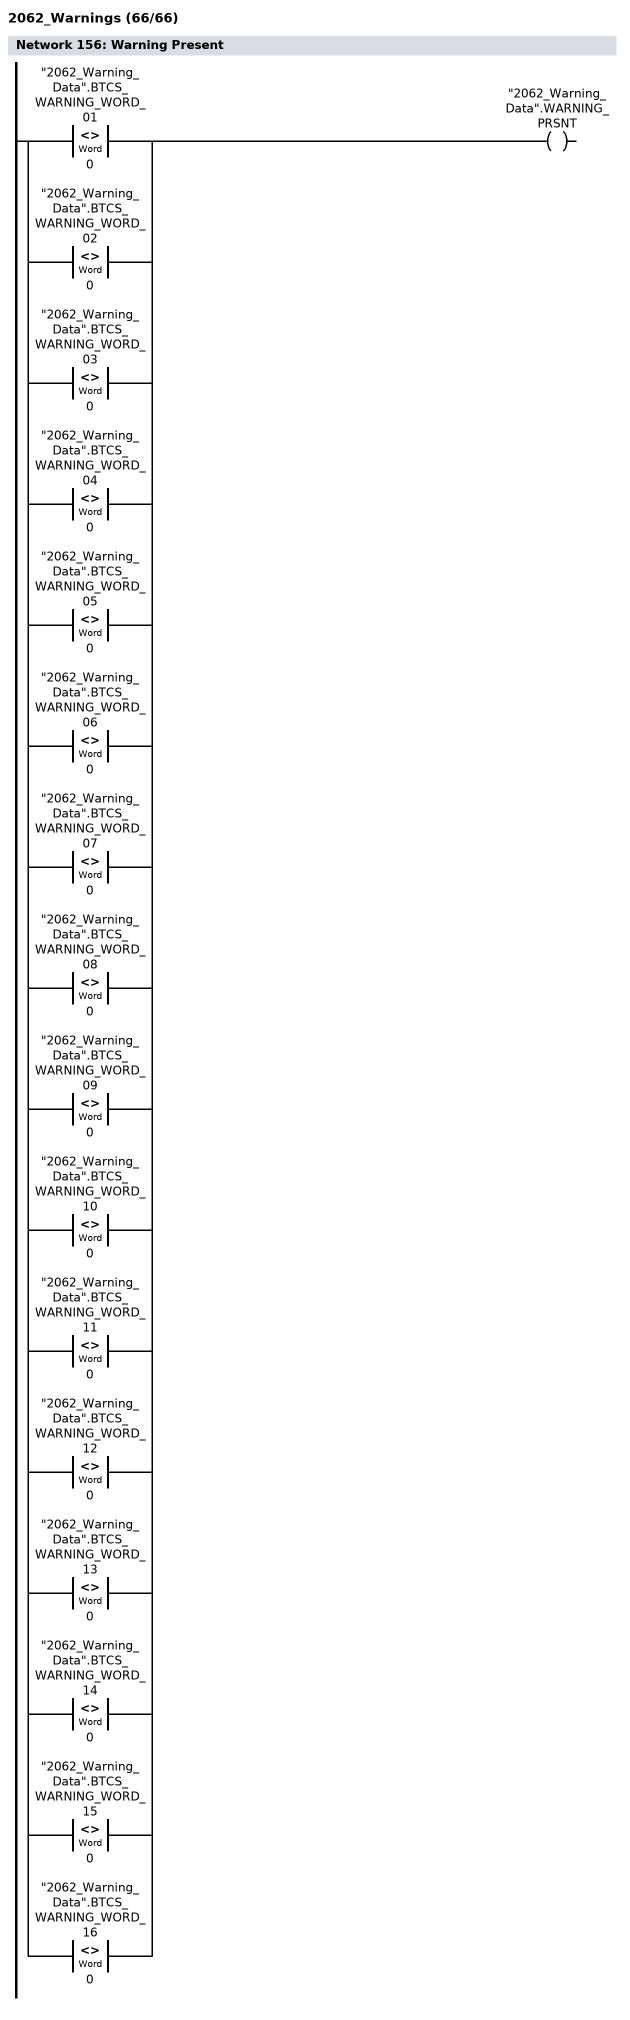
   RUNG wire#powerrail
      { S7_Templates := "SrcType := Word" } NE_Contact(in1 := "2062_Warning_Data".BTCS_WARNING_WORD_01, in2 := 0)
      wire#w1
      Coil( "2062_Warning_Data".WARNING_PRSNT )
   END_RUNG
   RUNG wire#powerrail
      { S7_Templates := "SrcType := Word" } NE_Contact(in1 := "2062_Warning_Data".BTCS_WARNING_WORD_02, in2 := 0)
   END_RUNG wire#w1
   RUNG wire#powerrail
      { S7_Templates := "SrcType := Word" } NE_Contact(in1 := "2062_Warning_Data".BTCS_WARNING_WORD_03, in2 := 0)
   END_RUNG wire#w1
   RUNG wire#powerrail
      { S7_Templates := "SrcType := Word" } NE_Contact(in1 := "2062_Warning_Data".BTCS_WARNING_WORD_04, in2 := 0)
   END_RUNG wire#w1
   RUNG wire#powerrail
      { S7_Templates := "SrcType := Word" } NE_Contact(in1 := "2062_Warning_Data".BTCS_WARNING_WORD_05, in2 := 0)
   END_RUNG wire#w1
   RUNG wire#powerrail
      { S7_Templates := "SrcType := Word" } NE_Contact(in1 := "2062_Warning_Data".BTCS_WARNING_WORD_06, in2 := 0)
   END_RUNG wire#w1
   RUNG wire#powerrail
      { S7_Templates := "SrcType := Word" } NE_Contact(in1 := "2062_Warning_Data".BTCS_WARNING_WORD_07, in2 := 0)
   END_RUNG wire#w1
   RUNG wire#powerrail
      { S7_Templates := "SrcType := Word" } NE_Contact(in1 := "2062_Warning_Data".BTCS_WARNING_WORD_08, in2 := 0)
   END_RUNG wire#w1
   RUNG wire#powerrail
      { S7_Templates := "SrcType := Word" } NE_Contact(in1 := "2062_Warning_Data".BTCS_WARNING_WORD_09, in2 := 0)
   END_RUNG wire#w1
   RUNG wire#powerrail
      { S7_Templates := "SrcType := Word" } NE_Contact(in1 := "2062_Warning_Data".BTCS_WARNING_WORD_10, in2 := 0)
   END_RUNG wire#w1
   RUNG wire#powerrail
      { S7_Templates := "SrcType := Word" } NE_Contact(in1 := "2062_Warning_Data".BTCS_WARNING_WORD_11, in2 := 0)
   END_RUNG wire#w1
   RUNG wire#powerrail
      { S7_Templates := "SrcType := Word" } NE_Contact(in1 := "2062_Warning_Data".BTCS_WARNING_WORD_12, in2 := 0)
   END_RUNG wire#w1
   RUNG wire#powerrail
      { S7_Templates := "SrcType := Word" } NE_Contact(in1 := "2062_Warning_Data".BTCS_WARNING_WORD_13, in2 := 0)
   END_RUNG wire#w1
   RUNG wire#powerrail
      { S7_Templates := "SrcType := Word" } NE_Contact(in1 := "2062_Warning_Data".BTCS_WARNING_WORD_14, in2 := 0)
   END_RUNG wire#w1
   RUNG wire#powerrail
      { S7_Templates := "SrcType := Word" } NE_Contact(in1 := "2062_Warning_Data".BTCS_WARNING_WORD_15, in2 := 0)
   END_RUNG wire#w1
   RUNG wire#powerrail
      { S7_Templates := "SrcType := Word" } NE_Contact(in1 := "2062_Warning_Data".BTCS_WARNING_WORD_16, in2 := 0)
   END_RUNG wire#w1
   // the same network as SCL:
   "2062_Warning_Data".WARNING_PRSNT := ("2062_Warning_Data".BTCS_WARNING_WORD_01 <> 0) OR ("2062_Warning_Data".BTCS_WARNING_WORD_02 <> 0) OR ("2062_Warning_Data".BTCS_WARNING_WORD_03 <> 0) OR ("2062_Warning_Data".BTCS_WARNING_WORD_04 <> 0) OR ("2062_Warning_Data".BTCS_WARNING_WORD_05 <> 0) OR ("2062_Warning_Data".BTCS_WARNING_WORD_06 <> 0) OR ("2062_Warning_Data".BTCS_WARNING_WORD_07 <> 0) OR ("2062_Warning_Data".BTCS_WARNING_WORD_08 <> 0) OR ("2062_Warning_Data".BTCS_WARNING_WORD_09 <> 0) OR ("2062_Warning_Data".BTCS_WARNING_WORD_10 <> 0) OR ("2062_Warning_Data".BTCS_WARNING_WORD_11 <> 0) OR ("2062_Warning_Data".BTCS_WARNING_WORD_12 <> 0) OR ("2062_Warning_Data".BTCS_WARNING_WORD_13 <> 0) OR ("2062_Warning_Data".BTCS_WARNING_WORD_14 <> 0) OR ("2062_Warning_Data".BTCS_WARNING_WORD_15 <> 0) OR ("2062_Warning_Data".BTCS_WARNING_WORD_16 <> 0);
END_REGION
END_FUNCTION

FUNCTION "2068_Sys_Status" : Void   // FC2068, LAD
TITLE = System Status
{ S7_Optimized_Access := 'TRUE' }
AUTHOR : JRS
VERSION : 0.1
// For the determination of specific system status information as required by the code
   VAR_TEMP
      RET_VAL_1 : Int;
      LOCAL_DATE_AND_TIME : DTL;
   END_VAR
   VAR_TEMP   // added for the SCL form of the ladder/FBD networks
      _w1 : Bool;
      _w2 : Bool;
      _w3 : Bool;
      _w4 : Bool;
   END_VAR
BEGIN

REGION Network 1: Port GTT Open Timer For Flow De-Bounce
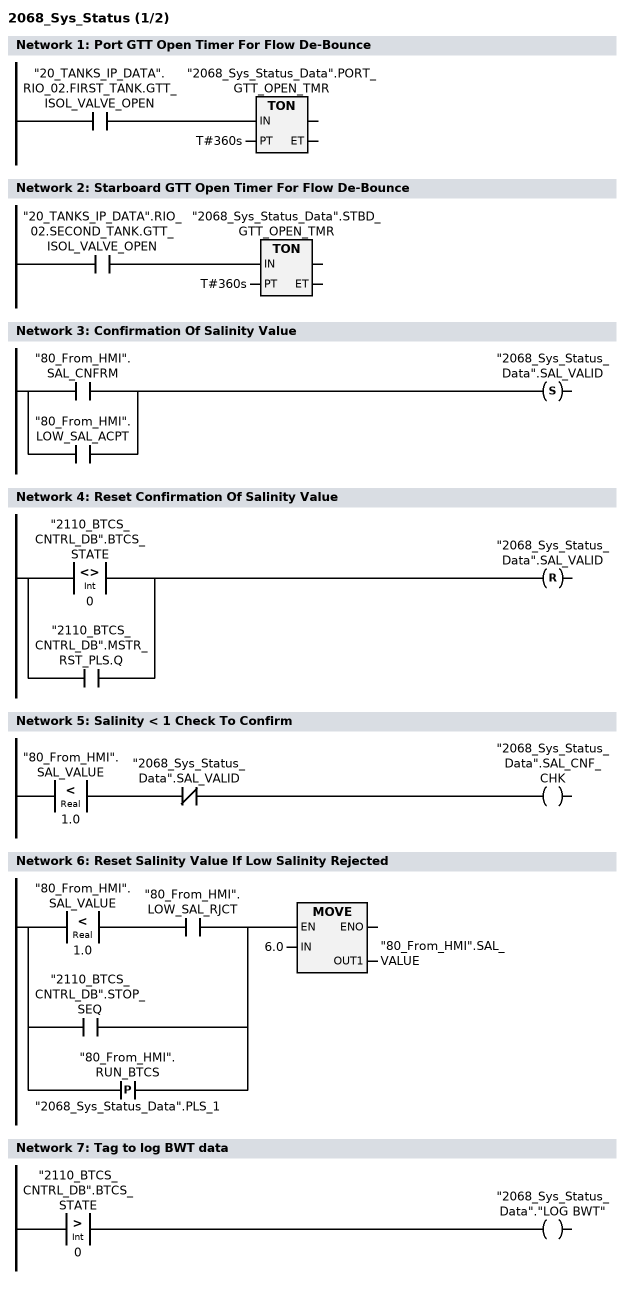
   "2068_Sys_Status_Data".PORT_GTT_OPEN_TMR.TON(IN := "20_TANKS_IP_DATA".RIO_02.FIRST_TANK.GTT_ISOL_VALVE_OPEN,
                           PT := T#360s);
END_REGION

REGION Network 2: Starboard GTT Open Timer For Flow De-Bounce
   "2068_Sys_Status_Data".STBD_GTT_OPEN_TMR.TON(IN := "20_TANKS_IP_DATA".RIO_02.SECOND_TANK.GTT_ISOL_VALVE_OPEN,
                           PT := T#360s);
END_REGION

REGION Network 3: Confirmation Of Salinity Value
   RUNG wire#powerrail
      Contact( "80_From_HMI".SAL_CNFRM )
      wire#w1
      S_Coil( "2068_Sys_Status_Data".SAL_VALID )
   END_RUNG
   RUNG wire#powerrail
      Contact( "80_From_HMI".LOW_SAL_ACPT )
   END_RUNG wire#w1
   // the same network as SCL:
   IF "80_From_HMI".SAL_CNFRM OR "80_From_HMI".LOW_SAL_ACPT THEN
       "2068_Sys_Status_Data".SAL_VALID := TRUE;
   END_IF;
END_REGION

REGION Network 4: Reset Confirmation Of Salinity Value
   RUNG wire#powerrail
      { S7_Templates := "SrcType := Int" } NE_Contact(in1 := "2110_BTCS_CNTRL_DB".BTCS_STATE, in2 := 0)
      wire#w1
      R_Coil( "2068_Sys_Status_Data".SAL_VALID )
   END_RUNG
   RUNG wire#powerrail
      Contact( "2110_BTCS_CNTRL_DB".MSTR_RST_PLS.Q )
   END_RUNG wire#w1
   // the same network as SCL:
   IF ("2110_BTCS_CNTRL_DB".BTCS_STATE <> 0) OR "2110_BTCS_CNTRL_DB".MSTR_RST_PLS.Q THEN
       "2068_Sys_Status_Data".SAL_VALID := FALSE;
   END_IF;
END_REGION

REGION Network 5: Salinity < 1 Check To Confirm
   RUNG wire#powerrail
      { S7_Templates := "SrcType := Real" } LT_Contact(in1 := "80_From_HMI".SAL_VALUE, in2 := 1.0)
      I_Contact( "2068_Sys_Status_Data".SAL_VALID )
      Coil( "2068_Sys_Status_Data".SAL_CNF_CHK )
   END_RUNG
   // the same network as SCL:
   "2068_Sys_Status_Data".SAL_CNF_CHK := ("80_From_HMI".SAL_VALUE < 1.0) AND NOT "2068_Sys_Status_Data".SAL_VALID;
END_REGION

REGION Network 6: Reset Salinity Value If Low Salinity Rejected
   RUNG wire#powerrail
      { S7_Templates := "SrcType := Real" } LT_Contact(in1 := "80_From_HMI".SAL_VALUE, in2 := 1.0)
      Contact( "80_From_HMI".LOW_SAL_RJCT )
      wire#w1
      Move(in := 6.0, out1 => "80_From_HMI".SAL_VALUE)
   END_RUNG
   RUNG wire#powerrail
      Contact( "2110_BTCS_CNTRL_DB".STOP_SEQ )
   END_RUNG wire#w1
   RUNG wire#powerrail
      P_Contact(operand := "80_From_HMI".RUN_BTCS, bit := "2068_Sys_Status_Data".PLS_1)
   END_RUNG wire#w1
   // the same network as SCL:
   #_w1 := "80_From_HMI".RUN_BTCS AND NOT "2068_Sys_Status_Data".PLS_1;   // rising edge of "80_From_HMI".RUN_BTCS
   "2068_Sys_Status_Data".PLS_1 := "80_From_HMI".RUN_BTCS;
   IF (("80_From_HMI".SAL_VALUE < 1.0) AND "80_From_HMI".LOW_SAL_RJCT) OR "2110_BTCS_CNTRL_DB".STOP_SEQ OR #_w1 THEN
       "80_From_HMI".SAL_VALUE := 6.0;
   END_IF;
END_REGION

REGION Network 7: Tag to log BWT data
   RUNG wire#powerrail
      { S7_Templates := "SrcType := Int" } GT_Contact(in1 := "2110_BTCS_CNTRL_DB".BTCS_STATE, in2 := 0)
      Coil( "2068_Sys_Status_Data"."LOG BWT" )
   END_RUNG
   // the same network as SCL:
   "2068_Sys_Status_Data"."LOG BWT" := "2110_BTCS_CNTRL_DB".BTCS_STATE > 0;
END_REGION

REGION Network 8
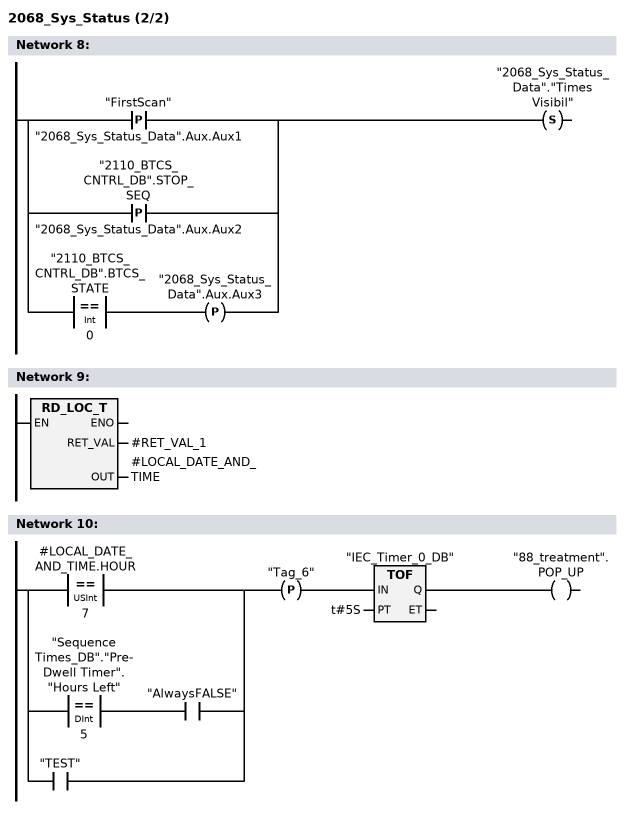
   RUNG wire#powerrail
      P_Contact(operand := "FirstScan", bit := "2068_Sys_Status_Data".Aux.Aux1)
      wire#w1
      S_Coil( "2068_Sys_Status_Data"."Times Visibil" )
   END_RUNG
   RUNG wire#powerrail
      P_Contact(operand := "2110_BTCS_CNTRL_DB".STOP_SEQ, bit := "2068_Sys_Status_Data".Aux.Aux2)
   END_RUNG wire#w1
   RUNG wire#powerrail
      { S7_Templates := "SrcType := Int" } EQ_Contact(in1 := "2110_BTCS_CNTRL_DB".BTCS_STATE, in2 := 0)
      P_Trig( "2068_Sys_Status_Data".Aux.Aux3 )
   END_RUNG wire#w1
   // the same network as SCL:
   #_w1 := "FirstScan" AND NOT "2068_Sys_Status_Data".Aux.Aux1;   // rising edge of "FirstScan"
   "2068_Sys_Status_Data".Aux.Aux1 := "FirstScan";
   #_w2 := "2110_BTCS_CNTRL_DB".STOP_SEQ AND NOT "2068_Sys_Status_Data".Aux.Aux2;   // rising edge of "2110_BTCS_CNTRL_DB".STOP_SEQ
   "2068_Sys_Status_Data".Aux.Aux2 := "2110_BTCS_CNTRL_DB".STOP_SEQ;
   #_w3 := "2110_BTCS_CNTRL_DB".BTCS_STATE = 0;
   #_w4 := #_w3 AND NOT "2068_Sys_Status_Data".Aux.Aux3;   // rising edge
   "2068_Sys_Status_Data".Aux.Aux3 := #_w3;
   IF #_w1 OR #_w2 OR #_w4 THEN "2068_Sys_Status_Data"."Times Visibil" := TRUE; END_IF;
END_REGION

REGION Network 9
   #RET_VAL_1 := RD_LOC_T(OUT => #LOCAL_DATE_AND_TIME);
END_REGION

REGION Network 10
   #_w1 := (#LOCAL_DATE_AND_TIME.HOUR = 7) OR (("Sequence Times_DB"."Pre-Dwell Timer"."Hours Left" = 5) AND "AlwaysFALSE") OR "TEST";
   #_w2 := #_w1 AND NOT "Tag_6";   // rising edge
   "Tag_6" := #_w1;
   "IEC_Timer_0_DB".TOF(IN := #_w2, PT := t#5S);
   "88_treatment".POP_UP := "IEC_Timer_0_DB".Q;
END_REGION
END_FUNCTION

// folder: 2000 - 2999 BTCS System/2100 - 2199 Automatic Sequencing

FUNCTION "2100_AUTO_SEQ" : Void   // FC2100, LAD
TITLE = Automatic Sequence
{ S7_Optimized_Access := 'TRUE' }
AUTHOR : JRS
VERSION : 0.1
// BTCS Automatic Sequence
   VAR_TEMP   // added for the SCL form of the ladder/FBD networks
      _w1 : Bool;
      _w2 : Bool;
      _w3 : Bool;
   END_VAR
BEGIN

REGION Network 1: Initialise Or Reset
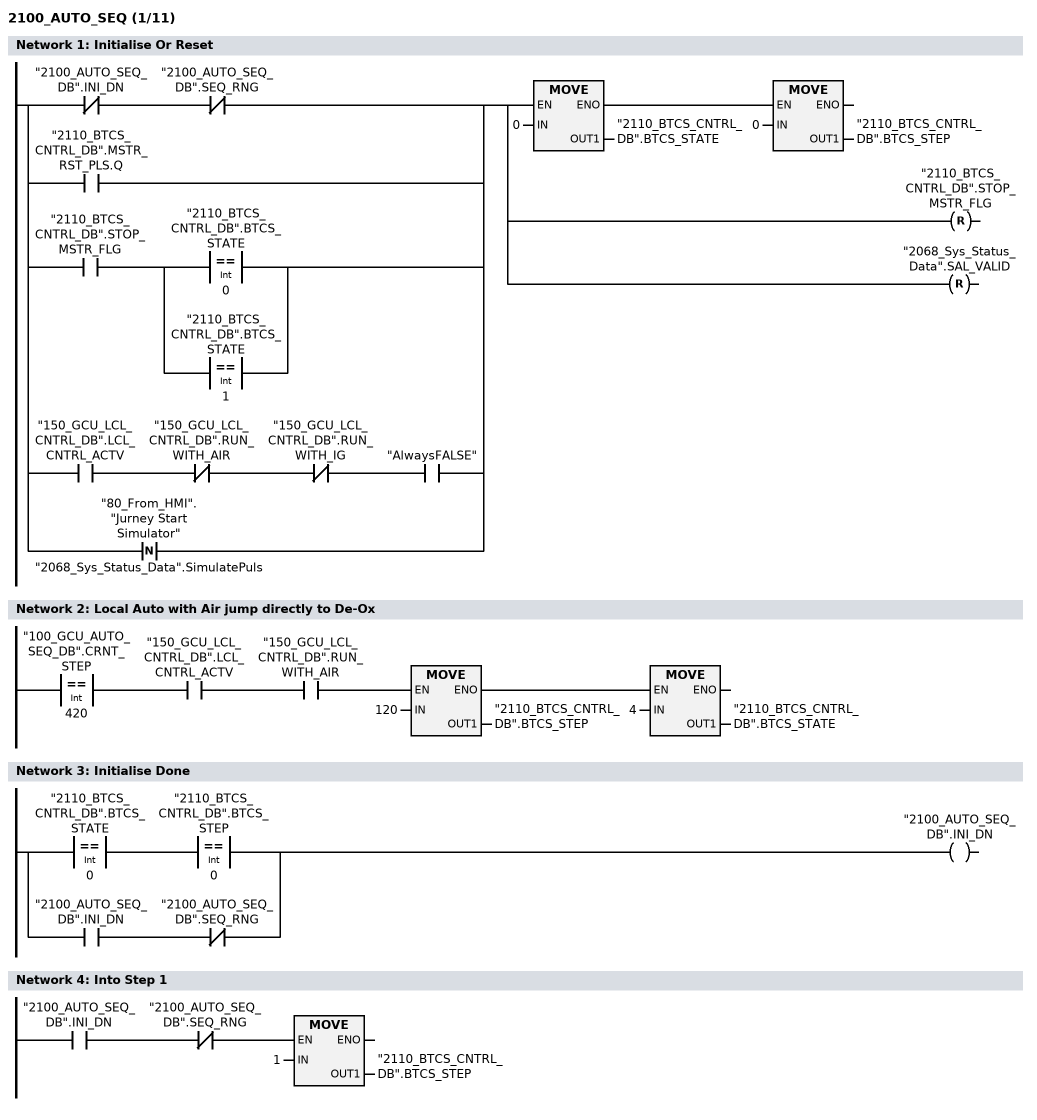
   RUNG wire#powerrail
      I_Contact( "2100_AUTO_SEQ_DB".INI_DN )
      I_Contact( "2100_AUTO_SEQ_DB".SEQ_RNG )
      wire#w1
      Move(in := 0, out1 => "2110_BTCS_CNTRL_DB".BTCS_STATE)
      Move(in := 0, out1 => "2110_BTCS_CNTRL_DB".BTCS_STEP)
   END_RUNG
   RUNG wire#powerrail
      Contact( "2110_BTCS_CNTRL_DB".MSTR_RST_PLS.Q )
   END_RUNG wire#w1
   RUNG wire#powerrail
      Contact( "2110_BTCS_CNTRL_DB".STOP_MSTR_FLG )
      wire#w2
      { S7_Templates := "SrcType := Int" } EQ_Contact(in1 := "2110_BTCS_CNTRL_DB".BTCS_STATE, in2 := 0)
   END_RUNG wire#w1
   RUNG wire#w2
      { S7_Templates := "SrcType := Int" } EQ_Contact(in1 := "2110_BTCS_CNTRL_DB".BTCS_STATE, in2 := 1)
   END_RUNG wire#w1
   RUNG wire#powerrail
      Contact( "150_GCU_LCL_CNTRL_DB".LCL_CNTRL_ACTV )
      I_Contact( "150_GCU_LCL_CNTRL_DB".RUN_WITH_AIR )
      I_Contact( "150_GCU_LCL_CNTRL_DB".RUN_WITH_IG )
      Contact( "AlwaysFALSE" )
   END_RUNG wire#w1
   RUNG wire#powerrail
      N_Contact(operand := "80_From_HMI"."Jurney Start Simulator", bit := "2068_Sys_Status_Data".SimulatePuls)
   END_RUNG wire#w1
   RUNG wire#w1
      R_Coil( "2110_BTCS_CNTRL_DB".STOP_MSTR_FLG )
   END_RUNG
   RUNG wire#w1
      R_Coil( "2068_Sys_Status_Data".SAL_VALID )
   END_RUNG
   // the same network as SCL:
   #_w1 := NOT "80_From_HMI"."Jurney Start Simulator" AND "2068_Sys_Status_Data".SimulatePuls;   // falling edge of "80_From_HMI"."Jurney Start Simulator"
   "2068_Sys_Status_Data".SimulatePuls := "80_From_HMI"."Jurney Start Simulator";
   #_w2 := (NOT "2100_AUTO_SEQ_DB".INI_DN AND NOT "2100_AUTO_SEQ_DB".SEQ_RNG) OR "2110_BTCS_CNTRL_DB".MSTR_RST_PLS.Q OR ("2110_BTCS_CNTRL_DB".STOP_MSTR_FLG AND (("2110_BTCS_CNTRL_DB".BTCS_STATE = 0) OR ("2110_BTCS_CNTRL_DB".BTCS_STATE = 1))) OR ("150_GCU_LCL_CNTRL_DB".LCL_CNTRL_ACTV AND NOT "150_GCU_LCL_CNTRL_DB".RUN_WITH_AIR AND NOT "150_GCU_LCL_CNTRL_DB".RUN_WITH_IG AND "AlwaysFALSE") OR #_w1;
   #_w3 := (NOT "2100_AUTO_SEQ_DB".INI_DN AND NOT "2100_AUTO_SEQ_DB".SEQ_RNG) OR "2110_BTCS_CNTRL_DB".MSTR_RST_PLS.Q OR ("2110_BTCS_CNTRL_DB".STOP_MSTR_FLG AND (("2110_BTCS_CNTRL_DB".BTCS_STATE = 0) OR ("2110_BTCS_CNTRL_DB".BTCS_STATE = 1))) OR ("150_GCU_LCL_CNTRL_DB".LCL_CNTRL_ACTV AND NOT "150_GCU_LCL_CNTRL_DB".RUN_WITH_AIR AND NOT "150_GCU_LCL_CNTRL_DB".RUN_WITH_IG AND "AlwaysFALSE") OR #_w1;
   IF #_w3 THEN
       "2110_BTCS_CNTRL_DB".BTCS_STATE := 0;
       "2110_BTCS_CNTRL_DB".BTCS_STEP := 0;
   END_IF;
   IF #_w2 THEN
       "2110_BTCS_CNTRL_DB".STOP_MSTR_FLG := FALSE;
       "2068_Sys_Status_Data".SAL_VALID := FALSE;
   END_IF;
END_REGION

REGION Network 2: Local Auto with Air jump directly to De-Ox
   RUNG wire#powerrail
      { S7_Templates := "SrcType := Int" } EQ_Contact(in1 := "100_GCU_AUTO_SEQ_DB".CRNT_STEP, in2 := 420)
      Contact( "150_GCU_LCL_CNTRL_DB".LCL_CNTRL_ACTV )
      Contact( "150_GCU_LCL_CNTRL_DB".RUN_WITH_AIR )
      Move(in := 120, out1 => "2110_BTCS_CNTRL_DB".BTCS_STEP)
      Move(in := 4, out1 => "2110_BTCS_CNTRL_DB".BTCS_STATE)
   END_RUNG
   // the same network as SCL:
   IF ("100_GCU_AUTO_SEQ_DB".CRNT_STEP = 420) AND "150_GCU_LCL_CNTRL_DB".LCL_CNTRL_ACTV AND "150_GCU_LCL_CNTRL_DB".RUN_WITH_AIR THEN
       "2110_BTCS_CNTRL_DB".BTCS_STEP := 120;
       "2110_BTCS_CNTRL_DB".BTCS_STATE := 4;
   END_IF;
END_REGION

REGION Network 3: Initialise Done
   RUNG wire#powerrail
      { S7_Templates := "SrcType := Int" } EQ_Contact(in1 := "2110_BTCS_CNTRL_DB".BTCS_STATE, in2 := 0)
      { S7_Templates := "SrcType := Int" } EQ_Contact(in1 := "2110_BTCS_CNTRL_DB".BTCS_STEP, in2 := 0)
      wire#w1
      Coil( "2100_AUTO_SEQ_DB".INI_DN )
   END_RUNG
   RUNG wire#powerrail
      Contact( "2100_AUTO_SEQ_DB".INI_DN )
      I_Contact( "2100_AUTO_SEQ_DB".SEQ_RNG )
   END_RUNG wire#w1
   // the same network as SCL:
   "2100_AUTO_SEQ_DB".INI_DN := (("2110_BTCS_CNTRL_DB".BTCS_STATE = 0) AND ("2110_BTCS_CNTRL_DB".BTCS_STEP = 0)) OR ("2100_AUTO_SEQ_DB".INI_DN AND NOT "2100_AUTO_SEQ_DB".SEQ_RNG);
END_REGION

REGION Network 4: Into Step 1
   RUNG wire#powerrail
      Contact( "2100_AUTO_SEQ_DB".INI_DN )
      I_Contact( "2100_AUTO_SEQ_DB".SEQ_RNG )
      Move(in := 1, out1 => "2110_BTCS_CNTRL_DB".BTCS_STEP)
   END_RUNG
   // the same network as SCL:
   IF "2100_AUTO_SEQ_DB".INI_DN AND NOT "2100_AUTO_SEQ_DB".SEQ_RNG THEN
       "2110_BTCS_CNTRL_DB".BTCS_STEP := 1;
   END_IF;
END_REGION

REGION Network 5: Step 1 = Wait For Accept & Launch (Times & Salinity Must Be Valid)
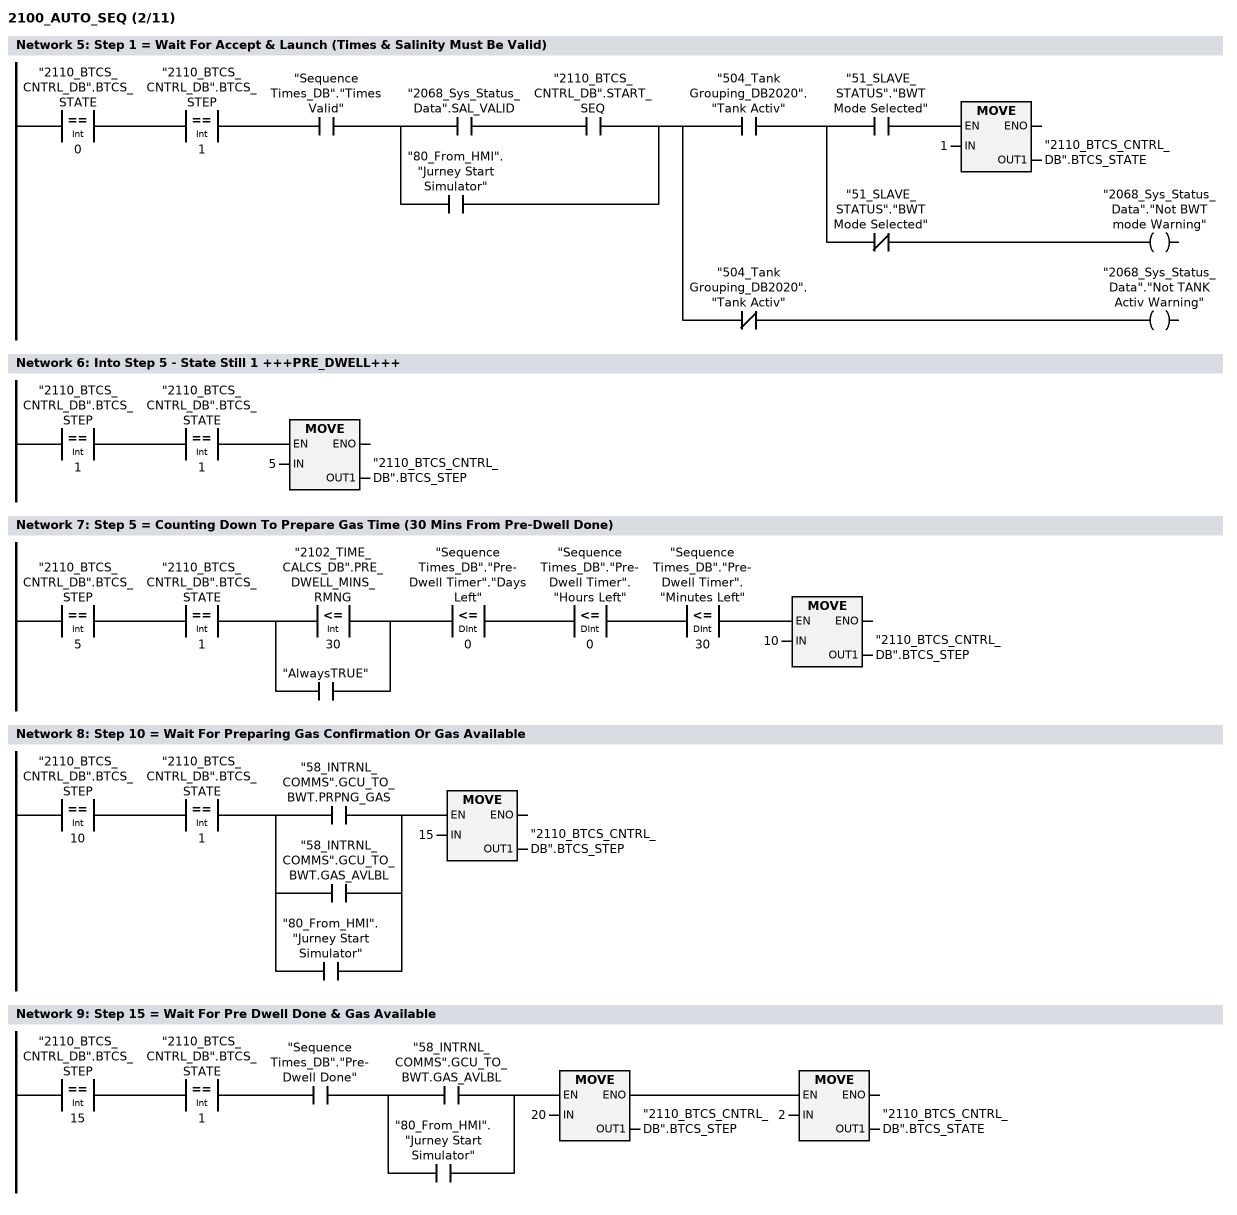
   RUNG wire#powerrail
      { S7_Templates := "SrcType := Int" } EQ_Contact(in1 := "2110_BTCS_CNTRL_DB".BTCS_STATE, in2 := 0)
      { S7_Templates := "SrcType := Int" } EQ_Contact(in1 := "2110_BTCS_CNTRL_DB".BTCS_STEP, in2 := 1)
      Contact( "Sequence Times_DB"."Times Valid" )
      wire#w1
      Contact( "2068_Sys_Status_Data".SAL_VALID )
      Contact( "2110_BTCS_CNTRL_DB".START_SEQ )
      wire#w2
      Contact( "504_Tank Grouping_DB2020"."Tank Activ" )
      wire#w3
      Contact( "51_SLAVE_STATUS"."BWT Mode Selected" )
      Move(in := 1, out1 => "2110_BTCS_CNTRL_DB".BTCS_STATE)
   END_RUNG
   RUNG wire#w1
      Contact( "80_From_HMI"."Jurney Start Simulator" )
   END_RUNG wire#w2
   RUNG wire#w3
      I_Contact( "51_SLAVE_STATUS"."BWT Mode Selected" )
      Coil( "2068_Sys_Status_Data"."Not BWT mode Warning" )
   END_RUNG
   RUNG wire#w2
      I_Contact( "504_Tank Grouping_DB2020"."Tank Activ" )
      Coil( "2068_Sys_Status_Data"."Not TANK Activ Warning" )
   END_RUNG
   // the same network as SCL:
   #_w1 := ("2110_BTCS_CNTRL_DB".BTCS_STATE = 0) AND ("2110_BTCS_CNTRL_DB".BTCS_STEP = 1) AND "Sequence Times_DB"."Times Valid" AND (("2068_Sys_Status_Data".SAL_VALID AND "2110_BTCS_CNTRL_DB".START_SEQ) OR "80_From_HMI"."Jurney Start Simulator");
   #_w2 := #_w1 AND "504_Tank Grouping_DB2020"."Tank Activ";
   IF #_w2 AND "51_SLAVE_STATUS"."BWT Mode Selected" THEN "2110_BTCS_CNTRL_DB".BTCS_STATE := 1; END_IF;
   "2068_Sys_Status_Data"."Not BWT mode Warning" := #_w2 AND NOT "51_SLAVE_STATUS"."BWT Mode Selected";
   "2068_Sys_Status_Data"."Not TANK Activ Warning" := #_w1 AND NOT "504_Tank Grouping_DB2020"."Tank Activ";
END_REGION

REGION Network 6: Into Step 5 - State Still 1 +++PRE_DWELL+++
   RUNG wire#powerrail
      { S7_Templates := "SrcType := Int" } EQ_Contact(in1 := "2110_BTCS_CNTRL_DB".BTCS_STEP, in2 := 1)
      { S7_Templates := "SrcType := Int" } EQ_Contact(in1 := "2110_BTCS_CNTRL_DB".BTCS_STATE, in2 := 1)
      Move(in := 5, out1 => "2110_BTCS_CNTRL_DB".BTCS_STEP)
   END_RUNG
   // the same network as SCL:
   IF ("2110_BTCS_CNTRL_DB".BTCS_STEP = 1) AND ("2110_BTCS_CNTRL_DB".BTCS_STATE = 1) THEN
       "2110_BTCS_CNTRL_DB".BTCS_STEP := 5;
   END_IF;
END_REGION

REGION Network 7: Step 5 = Counting Down To Prepare Gas Time (30 Mins From Pre-Dwell Done)
   RUNG wire#powerrail
      { S7_Templates := "SrcType := Int" } EQ_Contact(in1 := "2110_BTCS_CNTRL_DB".BTCS_STEP, in2 := 5)
      { S7_Templates := "SrcType := Int" } EQ_Contact(in1 := "2110_BTCS_CNTRL_DB".BTCS_STATE, in2 := 1)
      wire#w1
      { S7_Templates := "SrcType := Int" } LE_Contact(in1 := "2102_TIME_CALCS_DB".PRE_DWELL_MINS_RMNG, in2 := 30)
      wire#w2
      { S7_Templates := "SrcType := DInt" } LE_Contact(in1 := "Sequence Times_DB"."Pre-Dwell Timer"."Days Left", in2 := 0)
      { S7_Templates := "SrcType := DInt" } LE_Contact(in1 := "Sequence Times_DB"."Pre-Dwell Timer"."Hours Left", in2 := 0)
      { S7_Templates := "SrcType := DInt" } LE_Contact(in1 := "Sequence Times_DB"."Pre-Dwell Timer"."Minutes Left", in2 := 30)
      Move(in := 10, out1 => "2110_BTCS_CNTRL_DB".BTCS_STEP)
   END_RUNG
   RUNG wire#w1
      Contact( "AlwaysTRUE" )
   END_RUNG wire#w2
   // the same network as SCL:
   IF ("2110_BTCS_CNTRL_DB".BTCS_STEP = 5) AND ("2110_BTCS_CNTRL_DB".BTCS_STATE = 1) AND (("2102_TIME_CALCS_DB".PRE_DWELL_MINS_RMNG <= 30) OR "AlwaysTRUE") AND ("Sequence Times_DB"."Pre-Dwell Timer"."Days Left" <= 0) AND ("Sequence Times_DB"."Pre-Dwell Timer"."Hours Left" <= 0) AND ("Sequence Times_DB"."Pre-Dwell Timer"."Minutes Left" <= 30) THEN
       "2110_BTCS_CNTRL_DB".BTCS_STEP := 10;
   END_IF;
END_REGION

REGION Network 8: Step 10 = Wait For Preparing Gas Confirmation Or Gas Available
   RUNG wire#powerrail
      { S7_Templates := "SrcType := Int" } EQ_Contact(in1 := "2110_BTCS_CNTRL_DB".BTCS_STEP, in2 := 10)
      { S7_Templates := "SrcType := Int" } EQ_Contact(in1 := "2110_BTCS_CNTRL_DB".BTCS_STATE, in2 := 1)
      wire#w1
      Contact( "58_INTRNL_COMMS".GCU_TO_BWT.PRPNG_GAS )
      wire#w2
      Move(in := 15, out1 => "2110_BTCS_CNTRL_DB".BTCS_STEP)
   END_RUNG
   RUNG wire#w1
      Contact( "58_INTRNL_COMMS".GCU_TO_BWT.GAS_AVLBL )
   END_RUNG wire#w2
   RUNG wire#w1
      Contact( "80_From_HMI"."Jurney Start Simulator" )
   END_RUNG wire#w2
   // the same network as SCL:
   IF ("2110_BTCS_CNTRL_DB".BTCS_STEP = 10) AND ("2110_BTCS_CNTRL_DB".BTCS_STATE = 1) AND ("58_INTRNL_COMMS".GCU_TO_BWT.PRPNG_GAS OR "58_INTRNL_COMMS".GCU_TO_BWT.GAS_AVLBL OR "80_From_HMI"."Jurney Start Simulator") THEN
       "2110_BTCS_CNTRL_DB".BTCS_STEP := 15;
   END_IF;
END_REGION

REGION Network 9: Step 15 = Wait For Pre Dwell Done & Gas Available
   RUNG wire#powerrail
      { S7_Templates := "SrcType := Int" } EQ_Contact(in1 := "2110_BTCS_CNTRL_DB".BTCS_STEP, in2 := 15)
      { S7_Templates := "SrcType := Int" } EQ_Contact(in1 := "2110_BTCS_CNTRL_DB".BTCS_STATE, in2 := 1)
      Contact( "Sequence Times_DB"."Pre-Dwell Done" )
      wire#w1
      Contact( "58_INTRNL_COMMS".GCU_TO_BWT.GAS_AVLBL )
      wire#w2
      Move(in := 20, out1 => "2110_BTCS_CNTRL_DB".BTCS_STEP)
      Move(in := 2, out1 => "2110_BTCS_CNTRL_DB".BTCS_STATE)
   END_RUNG
   RUNG wire#w1
      Contact( "80_From_HMI"."Jurney Start Simulator" )
   END_RUNG wire#w2
   // the same network as SCL:
   #_w1 := ("2110_BTCS_CNTRL_DB".BTCS_STEP = 15) AND ("2110_BTCS_CNTRL_DB".BTCS_STATE = 1) AND "Sequence Times_DB"."Pre-Dwell Done" AND ("58_INTRNL_COMMS".GCU_TO_BWT.GAS_AVLBL OR "80_From_HMI"."Jurney Start Simulator");
   IF #_w1 THEN
       "2110_BTCS_CNTRL_DB".BTCS_STEP := 20;
       "2110_BTCS_CNTRL_DB".BTCS_STATE := 2;
   END_IF;
END_REGION

REGION Network 10: Step 20 = Close All Activated Tank Vent Valves +++DE_OX+++
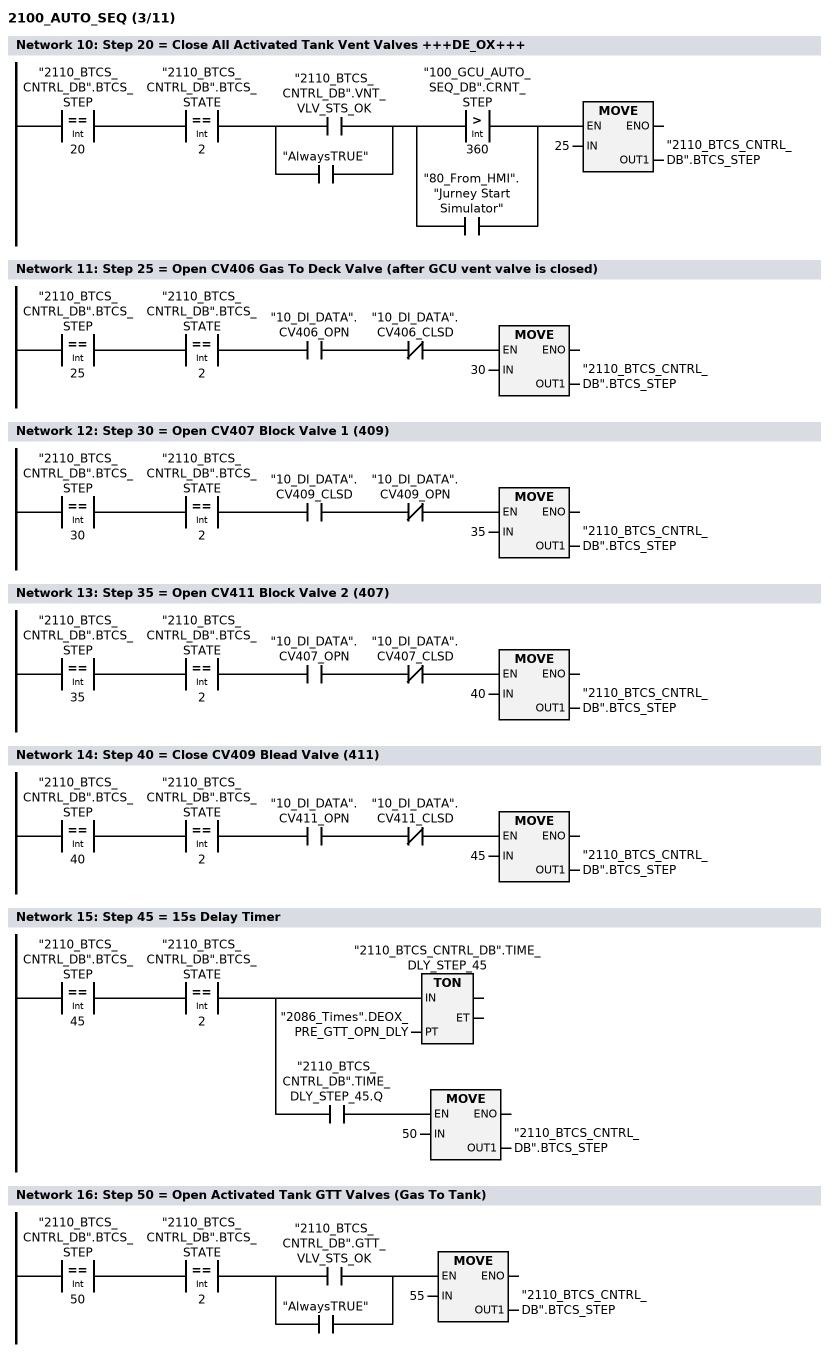
   RUNG wire#powerrail
      { S7_Templates := "SrcType := Int" } EQ_Contact(in1 := "2110_BTCS_CNTRL_DB".BTCS_STEP, in2 := 20)
      { S7_Templates := "SrcType := Int" } EQ_Contact(in1 := "2110_BTCS_CNTRL_DB".BTCS_STATE, in2 := 2)
      wire#w1
      Contact( "2110_BTCS_CNTRL_DB".VNT_VLV_STS_OK )
      wire#w2
      { S7_Templates := "SrcType := Int" } GT_Contact(in1 := "100_GCU_AUTO_SEQ_DB".CRNT_STEP, in2 := 360)
      wire#w3
      Move(in := 25, out1 => "2110_BTCS_CNTRL_DB".BTCS_STEP)
   END_RUNG
   RUNG wire#w1
      Contact( "AlwaysTRUE" )
   END_RUNG wire#w2
   RUNG wire#w2
      Contact( "80_From_HMI"."Jurney Start Simulator" )
   END_RUNG wire#w3
   // the same network as SCL:
   IF ("2110_BTCS_CNTRL_DB".BTCS_STEP = 20) AND ("2110_BTCS_CNTRL_DB".BTCS_STATE = 2) AND ("2110_BTCS_CNTRL_DB".VNT_VLV_STS_OK OR "AlwaysTRUE") AND (("100_GCU_AUTO_SEQ_DB".CRNT_STEP > 360) OR "80_From_HMI"."Jurney Start Simulator") THEN
       "2110_BTCS_CNTRL_DB".BTCS_STEP := 25;
   END_IF;
END_REGION

REGION Network 11: Step 25 = Open CV406 Gas To Deck Valve (after GCU vent valve is closed)
   RUNG wire#powerrail
      { S7_Templates := "SrcType := Int" } EQ_Contact(in1 := "2110_BTCS_CNTRL_DB".BTCS_STEP, in2 := 25)
      { S7_Templates := "SrcType := Int" } EQ_Contact(in1 := "2110_BTCS_CNTRL_DB".BTCS_STATE, in2 := 2)
      Contact( "10_DI_DATA".CV406_OPN )
      I_Contact( "10_DI_DATA".CV406_CLSD )
      Move(in := 30, out1 => "2110_BTCS_CNTRL_DB".BTCS_STEP)
   END_RUNG
   // the same network as SCL:
   IF ("2110_BTCS_CNTRL_DB".BTCS_STEP = 25) AND ("2110_BTCS_CNTRL_DB".BTCS_STATE = 2) AND "10_DI_DATA".CV406_OPN AND NOT "10_DI_DATA".CV406_CLSD THEN
       "2110_BTCS_CNTRL_DB".BTCS_STEP := 30;
   END_IF;
END_REGION

REGION Network 12: Step 30 = Open CV407 Block Valve 1 (409)
   RUNG wire#powerrail
      { S7_Templates := "SrcType := Int" } EQ_Contact(in1 := "2110_BTCS_CNTRL_DB".BTCS_STEP, in2 := 30)
      { S7_Templates := "SrcType := Int" } EQ_Contact(in1 := "2110_BTCS_CNTRL_DB".BTCS_STATE, in2 := 2)
      Contact( "10_DI_DATA".CV409_CLSD )
      I_Contact( "10_DI_DATA".CV409_OPN )
      Move(in := 35, out1 => "2110_BTCS_CNTRL_DB".BTCS_STEP)
   END_RUNG
   // the same network as SCL:
   IF ("2110_BTCS_CNTRL_DB".BTCS_STEP = 30) AND ("2110_BTCS_CNTRL_DB".BTCS_STATE = 2) AND "10_DI_DATA".CV409_CLSD AND NOT "10_DI_DATA".CV409_OPN THEN
       "2110_BTCS_CNTRL_DB".BTCS_STEP := 35;
   END_IF;
END_REGION

REGION Network 13: Step 35 = Open CV411 Block Valve 2 (407)
   RUNG wire#powerrail
      { S7_Templates := "SrcType := Int" } EQ_Contact(in1 := "2110_BTCS_CNTRL_DB".BTCS_STEP, in2 := 35)
      { S7_Templates := "SrcType := Int" } EQ_Contact(in1 := "2110_BTCS_CNTRL_DB".BTCS_STATE, in2 := 2)
      Contact( "10_DI_DATA".CV407_OPN )
      I_Contact( "10_DI_DATA".CV407_CLSD )
      Move(in := 40, out1 => "2110_BTCS_CNTRL_DB".BTCS_STEP)
   END_RUNG
   // the same network as SCL:
   IF ("2110_BTCS_CNTRL_DB".BTCS_STEP = 35) AND ("2110_BTCS_CNTRL_DB".BTCS_STATE = 2) AND "10_DI_DATA".CV407_OPN AND NOT "10_DI_DATA".CV407_CLSD THEN
       "2110_BTCS_CNTRL_DB".BTCS_STEP := 40;
   END_IF;
END_REGION

REGION Network 14: Step 40 = Close CV409 Blead Valve (411)
   RUNG wire#powerrail
      { S7_Templates := "SrcType := Int" } EQ_Contact(in1 := "2110_BTCS_CNTRL_DB".BTCS_STEP, in2 := 40)
      { S7_Templates := "SrcType := Int" } EQ_Contact(in1 := "2110_BTCS_CNTRL_DB".BTCS_STATE, in2 := 2)
      Contact( "10_DI_DATA".CV411_OPN )
      I_Contact( "10_DI_DATA".CV411_CLSD )
      Move(in := 45, out1 => "2110_BTCS_CNTRL_DB".BTCS_STEP)
   END_RUNG
   // the same network as SCL:
   IF ("2110_BTCS_CNTRL_DB".BTCS_STEP = 40) AND ("2110_BTCS_CNTRL_DB".BTCS_STATE = 2) AND "10_DI_DATA".CV411_OPN AND NOT "10_DI_DATA".CV411_CLSD THEN
       "2110_BTCS_CNTRL_DB".BTCS_STEP := 45;
   END_IF;
END_REGION

REGION Network 15: Step 45 = 15s Delay Timer
   #_w1 := ("2110_BTCS_CNTRL_DB".BTCS_STEP = 45) AND ("2110_BTCS_CNTRL_DB".BTCS_STATE = 2);
   "2110_BTCS_CNTRL_DB".TIME_DLY_STEP_45.TON(IN := #_w1, PT := "2086_Times".DEOX_PRE_GTT_OPN_DLY);
   IF #_w1 AND "2110_BTCS_CNTRL_DB".TIME_DLY_STEP_45.Q THEN "2110_BTCS_CNTRL_DB".BTCS_STEP := 50; END_IF;
END_REGION

REGION Network 16: Step 50 = Open Activated Tank GTT Valves (Gas To Tank)
   RUNG wire#powerrail
      { S7_Templates := "SrcType := Int" } EQ_Contact(in1 := "2110_BTCS_CNTRL_DB".BTCS_STEP, in2 := 50)
      { S7_Templates := "SrcType := Int" } EQ_Contact(in1 := "2110_BTCS_CNTRL_DB".BTCS_STATE, in2 := 2)
      wire#w1
      Contact( "2110_BTCS_CNTRL_DB".GTT_VLV_STS_OK )
      wire#w2
      Move(in := 55, out1 => "2110_BTCS_CNTRL_DB".BTCS_STEP)
   END_RUNG
   RUNG wire#w1
      Contact( "AlwaysTRUE" )
   END_RUNG wire#w2
   // the same network as SCL:
   IF ("2110_BTCS_CNTRL_DB".BTCS_STEP = 50) AND ("2110_BTCS_CNTRL_DB".BTCS_STATE = 2) AND ("2110_BTCS_CNTRL_DB".GTT_VLV_STS_OK OR "AlwaysTRUE") THEN
       "2110_BTCS_CNTRL_DB".BTCS_STEP := 55;
   END_IF;
END_REGION

REGION Network 17: Step 55 = Wait For O2 <= SP For Active Tanks For 1 minute